// TIA Portal project "Canarias Skills" (V17)
// Prueba de periferia descentralizada ET 200SP

(* hardware
DEVICE "S7-1200 station_1"  S7-1200 Station
   slot 0: "Rack_0"  S7-1200 Rack  Rack  V1.0
   slot 1: "PLC"  CPU 1215C AC/DC/Rly  6ES7 215-1BG40-0XB0  V4.5
DEVICE "GSD device_1"  GSD.Device.PN
   slot 0: "Rack"  Rack  V1.0
   slot 0: "MASTER IO-Link"  AL1100  AL1100
      slot 0: "AL1100"  AL1100
      slot 1: "X1"  X1
         slot 1: "Port 1"  Port 1
         slot 2: "Port 2"  Port 2
      slot 1: "4 Ports_1"  4 Ports  AL1100
         slot 0: "IO-Link Master"  IO-Link Master
   slot 1: "Encoder"  IO-Link In  2 Byte + PQI
   slot 2: "PE"  Digital Input + PQI
   slot 3: "Capacitivo"  Digital Input + PQI
   slot 4: "Disabled_1"  Disabled
DEVICE "SINAMICS G_1"  Sinamics.Device
   slot 0: "	_0"  Rail  SinamicsG120SVecto
   slot 0: "DRIVE_cinta"  G120 CU250S-2 PN Vector  6SL3246-0BA22-1FA0  4.6
      slot 1: "PROFINET interface"  MDD-SinamicsG120-P
   slot 3: "PM240-2 IP20"  PM240-2 IP20  6SL3210-1PB13-8ULx  -
DEVICE "ET 200SP station_1"  ET 200SP-Station
   slot 0: "Rack_0"  Rack  6ES5 710-8MAx1
   slot 0: "IO device_1"  IM 155-6 PN HF  6ES7 155-6AU00-0CN0  V3.1
   slot 1: "DI 8x24VDC HF_1"  DI 8x24VDC HF  6ES7 131-6BF00-0CA0  V1.2
      slot 1: "DI 8x24VDC HF_1"  DI 8x24VDC HF
   slot 2: "DQ 8x24VDC/0.5A HF_1"  DQ 8x24VDC/0.5A HF  6ES7 132-6BF00-0CA0  V1.2
      slot 1: "DQ 8x24VDC/0.5A HF_1"  DQ 8x24VDC/0.5A HF
   slot 3: "Server module_1"  Server module  6ES7 193-6PA00-0AA0  V1.1
      slot 1: "Server module_1"  Server module
   slot 127: "BA 2xRJ45"  BA 2xRJ45  6ES7 193-6AR00-0AA0  V0.0
      slot 1: "Port_1"  X1 P1 R  6ES7 193-6AR00-0AA0  V0.0
      slot 2: "Port_2"  X1 P2 R  6ES7 193-6AR00-0AA0  V0.0
DEVICE "HMI"  KTP700 Basic PN
   slot 0: "HMI"  KTP700 Basic PN  6AV2 123-2GB03-0AX0  17.0.0.0
   slot 1: "HMI_RT_1"  KTP700 Basic PN  6AV2 123-2GB03-0AX0  17.0.0.0
   slot 5: "HMI.IE_CP_1"  PROFINET Interface  17.0.0.0
      slot 1: "PROFINET Interface_1"  PROFINET Interface
         slot 1: "Port_1"  Port
*)

// ===== PLC "PLC"  CPU 1215C AC/DC/Rly =====

VAR_GLOBAL   // PLC tag table "Default tag table"
   "System_Byte" AT %MB1 : Byte;
   "FirstScan" AT %M1.0 : Bool;
   "DiagStatusUpdate" AT %M1.1 : Bool;
   "AlwaysTRUE" AT %M1.2 : Bool;
   "AlwaysFALSE" AT %M1.3 : Bool;
   "Clock_Byte" AT %MB0 : Byte;
   "Clock_10Hz" AT %M0.0 : Bool;
   "Clock_5Hz" AT %M0.1 : Bool;
   "Clock_2.5Hz" AT %M0.2 : Bool;
   "Clock_2Hz" AT %M0.3 : Bool;
   "Clock_1.25Hz" AT %M0.4 : Bool;
   "Clock_1Hz" AT %M0.5 : Bool;
   "Clock_0.625Hz" AT %M0.6 : Bool;
   "Clock_0.5Hz" AT %M0.7 : Bool;
   "Tag_1" AT %Q256.7 : Bool;
   "Tag_2" AT %Q257.7 : Bool;
   "Tag_3" AT %I0.0 : Bool;
   "Tag_4" AT %Q0.0 : Bool;
   "Tag_5" AT %M100.0 : Bool;
END_VAR

VAR_GLOBAL   // PLC tag table "Tag table_1"
   "Encoder" AT %IW68 : Word;
   "Envase" AT %I2.0 : Bool;
   "Llenador_retroceder" AT %Q2.0 : Bool;
   "Llenador_avanzar" AT %Q2.2 : Bool;
   "Cargar_tapa_retroceder" AT %Q2.4 : Bool;
   "Cargar_tapa_avanzar" AT %Q2.6 : Bool;
   "Taponador_retroceder" AT %Q2.1 : Bool;
   "Taponador_avanzar" AT %Q2.5 : Bool;
   "Cargar_tapa_atras" AT %I3.0 : Bool;
   "Cargar_tapa_adelante" AT %I3.1 : Bool;
   "Taponador_atras" AT %I3.2 : Bool;
   "Taponador_adelante" AT %I3.3 : Bool;
   "Mando_driver_cinta" AT %QW256 : Word;
   "Consigna_driver_cinta" AT %QW258 : Word;
   "Estado_driver_cinta" AT %IW256 : Word;
   "Velocidad_cinta" AT %IW258 : Word;
   "R_distancia" AT %M210.0 : Bool;   // Borrar el contador de distancia de la cinta
   "PV_distancia" AT %MW212 : Word;   // Distancia que debe avanzar la cinta
   "Pulso_encoder" AT %I69.0 : Bool;   // Los pulsos del encoder marcan el avance de la cinta
   "PE" AT %I4.1 : Bool;   // Paro de energencia NC
   "CV_distancia" AT %MW214 : Word;   // Distancia que ha recorrido la cinta
   "Q_distancia" AT %M210.1 : Bool;   // Indica que la cinta recorrió la distancia programada
   "Alarmas" AT %MW100 : Word;   // Bits de alarma del HMI
   "ACK_alarmas" AT %MW102 : Word;   // Bits de reconocimiento de alarmas
END_VAR

DATA_BLOCK "Modbus Connect"   // DB1
{ S7_Optimized_Access := 'FALSE' }
VERSION : 0.1
   VAR
      Arduino_1 : Struct
         Configuration : TCON_IP_v4;
         Status : Word;
      END_STRUCT;
   END_VAR
BEGIN
   Arduino_1.Configuration.InterfaceId := 64;
   Arduino_1.Configuration.ID := 16#1;
   Arduino_1.Configuration.ActiveEstablished := TRUE;
   Arduino_1.Configuration.RemoteAddress.ADDR[4] := 200;
   Arduino_1.Configuration.RemoteAddress.ADDR[3] := 0;
   Arduino_1.Configuration.RemoteAddress.ADDR[2] := 168;
   Arduino_1.Configuration.RemoteAddress.ADDR[1] := 192;
   Arduino_1.Configuration.RemotePort := 502;
   Arduino_1.Configuration.LocalPort := 0;
END_DATA_BLOCK

DATA_BLOCK "Modbus Buffer"   // DB3
{ S7_Optimized_Access := 'FALSE' }
VERSION : 0.1
   VAR
      Datos : Array[0..100] of Word;
   END_VAR
BEGIN
END_DATA_BLOCK

DATA_BLOCK "Modo_automatico_DB"   // DB4
{ S7_Optimized_Access := 'TRUE' }
VERSION : 0.1
// stored: InstanceOfName Modo_automatico
"Modo_automatico"
BEGIN
END_DATA_BLOCK

DATA_BLOCK "Datos_maquina"   // DB5
{ S7_Optimized_Access := 'TRUE' }
VERSION : 0.1
   VAR RETAIN
      pp_mm : Int := 2;   // Pulsos de encoder por cada milímetro de avance de cinta
      Desviador_bloquear : Word := 0;   // Posición del desviador para bloquear pieza
      Desviador_rechazar : Word := 37;   // Posición del desviador para rechazar pieza
      Desviador_aceptar : Word := 82;   // Posición del desviador para aceptar pieza
      Distancia_inspeccion : Word := 50;   // Distancia en mm hasta el inspector
      Distancia_desviador : Word := 100;   // Distancia en mm hasta el desviador
      Distancia_llenadora : Word := 200;   // Distancia en mm hasta la llenadora
      Distancia_taponadora : Word := 300;   // Distancia en mm hasta la taponadora
      Distancia_salida : Word := 400;   // Distancia en mm hasta la salida de la cinta
      Cinta_en_espera : Word := 16#047E;   // Driver cinta listo y en espera
      Cinta_en_marcha : Word := 16#0C7F;   // Driver cinta en avance
      Consigna_cinta : Int := 8000;   // Consigna de velocidad de la cinta
      Freno_en_cinta : Word := 16#043F;   // Activar freno con rampa driver cinta
      Freno_en_cinta_rapido : Word := 16#043D;   // Activar freno rápìdo driver cinta
      Total_envasados : Word;   // Catidad de envases producidos
      Total_rechazados : Word;   // Cantidad de envases rechazados
   END_VAR
   VAR
      HMI_llenador_retroceder : Bool;   // Lo que sigue son maniobras en modo manual desde el HMI
      HMI_llenador_avanzar : Bool;
      HMI_cargar_tapa_retroceder : Bool;
      HMI_cargar_tapa_avanzar : Bool;
      HMI_taponar_retroceder : Bool;
      HMI_taponar_avanzar : Bool;
      HMI_desviador_bloquear : Bool;
      HMI_desviador_rechazar : Bool;
      HMI_desviador_aceptar : Bool;
      HMI_driver_listo : Bool;
      HMI_driver_acusar_fallo : Bool;   // Manobras en modo manual de la cinta
      HMI_driver_detener_rampa : Bool;
      HMI_driver_detener_freno : Bool;
      HMI_driver_marcha : Bool;
      HMI_marcha : Bool;   // Marcha desde el HMI
      HMI_paro : Bool;   // Paro desde el HMI
      HMI_reset : Bool;   // Reset desde el HMI
   END_VAR
   VAR RETAIN
      HMI_manual_automatico : Bool;   // Modo de operación desde el HMI
      Estado : Struct
         Esperando_marcha : Bool;
         En_marcha : Bool;
         En_paro : Bool;
         En_PE : Bool;
         Esperando_reset : Bool;
      END_STRUCT;
   END_VAR
   VAR
      Inspector : Struct
         Enviar : Bool;
         Recibir : Bool;
         Recibido_ok : Bool;
         Recibido_error : Bool;
      END_STRUCT;
   END_VAR
BEGIN
END_DATA_BLOCK

DATA_BLOCK "Paro_emergencia_DB"   // DB10
{ S7_Optimized_Access := 'TRUE' }
VERSION : 0.1
// stored: InstanceOfName Paro_emergencia
"Paro_emergencia"
BEGIN
END_DATA_BLOCK

DATA_BLOCK "Raspberry PI Buffer"   // DB13
{ S7_Optimized_Access := 'FALSE' }
VERSION : 0.1
   VAR
      Data_send : Array[0..100] of Char;
      Data_rcv : Array[0..29] of Char;
   END_VAR
BEGIN
   Data_send[9] := '"';
   Data_send[8] := 'd';
   Data_send[7] := 'n';
   Data_send[6] := 'a';
   Data_send[5] := 'm';
   Data_send[4] := 'm';
   Data_send[3] := 'o';
   Data_send[2] := 'c';
   Data_send[1] := '"';
   Data_send[0] := '{';
   Data_send[10] := ':';   // {Command=I} para inferir objeto
   Data_send[11] := '"';
   Data_send[12] := 'I';
   Data_send[13] := '"';
   Data_send[14] := '}';
END_DATA_BLOCK

// folder: System blocks/Program resources

DATA_BLOCK "Distancia"   // DB6
{ S7_Optimized_Access := 'TRUE' }
AUTHOR : Simatic
FAMILY : IEC
NAME : CNTR
VERSION : 1.0
// stored: InstanceOfName IEC_COUNTER
"IEC_COUNTER"
BEGIN
END_DATA_BLOCK

DATA_BLOCK "IEC_Timer_0_DB"   // DB7
{ S7_Optimized_Access := 'TRUE' }
AUTHOR : Simatic
FAMILY : IEC
NAME : IEC_TMR
VERSION : 1.0
// stored: InstanceOfName IEC_TIMER
"IEC_TIMER"
BEGIN
END_DATA_BLOCK

DATA_BLOCK "IEC_Timer_0_DB_1"   // DB8
{ S7_Optimized_Access := 'TRUE' }
AUTHOR : Simatic
FAMILY : IEC
NAME : IEC_TMR
VERSION : 1.0
// stored: InstanceOfName IEC_TIMER
"IEC_TIMER"
BEGIN
END_DATA_BLOCK

DATA_BLOCK "IEC_Timer_0_DB_2"   // DB9
{ S7_Optimized_Access := 'TRUE' }
AUTHOR : Simatic
FAMILY : IEC
NAME : IEC_TMR
VERSION : 1.0
// stored: InstanceOfName IEC_TIMER
"IEC_TIMER"
BEGIN
END_DATA_BLOCK

DATA_BLOCK "IEC_Timer_0_DB_3"   // DB11
{ S7_Optimized_Access := 'TRUE' }
AUTHOR : Simatic
FAMILY : IEC
NAME : IEC_TMR
VERSION : 1.0
// stored: InstanceOfName IEC_TIMER
"IEC_TIMER"
BEGIN
END_DATA_BLOCK

DATA_BLOCK "PLC_Receive_DB"   // DB15
{ S7_Optimized_Access := 'TRUE' }
AUTHOR : SIMATIC
FAMILY : MC7Plus
NAME : TC_IP_v4
VERSION : 1.0
// stored: InstanceOfName TCON_IP_v4
"TCON_IP_v4"
BEGIN
   ID := 3;
   InterfaceId := 64;
   LocalPort := 2000;
   RemotePort := 2000;
   ActiveEstablished := true;
   RemoteAddress.ADDR[1] := 192;
   RemoteAddress.ADDR[2] := 168;
   RemoteAddress.ADDR[4] := 241;
END_DATA_BLOCK

DATA_BLOCK "IEC_Timer_0_DB_4"   // DB16
{ S7_Optimized_Access := 'TRUE' }
AUTHOR : Simatic
FAMILY : IEC
NAME : IEC_TMR
VERSION : 1.0
// stored: InstanceOfName IEC_TIMER
"IEC_TIMER"
BEGIN
END_DATA_BLOCK

DATA_BLOCK "IEC_Timer_0_DB_5"   // DB17
{ S7_Optimized_Access := 'TRUE' }
AUTHOR : Simatic
FAMILY : IEC
NAME : IEC_TMR
VERSION : 1.0
// stored: InstanceOfName IEC_TIMER
"IEC_TIMER"
BEGIN
END_DATA_BLOCK

DATA_BLOCK "IEC_Timer_0_DB_6"   // DB18
{ S7_Optimized_Access := 'TRUE' }
AUTHOR : Simatic
FAMILY : IEC
NAME : IEC_TMR
VERSION : 1.0
// stored: InstanceOfName IEC_TIMER
"IEC_TIMER"
BEGIN
END_DATA_BLOCK

DATA_BLOCK "IEC_Timer_0_DB_7"   // DB19
{ S7_Optimized_Access := 'TRUE' }
AUTHOR : Simatic
FAMILY : IEC
NAME : IEC_TMR
VERSION : 1.0
// stored: InstanceOfName IEC_TIMER
"IEC_TIMER"
BEGIN
END_DATA_BLOCK

// folder: (top level)

FUNCTION_BLOCK "Paro_emergencia"   // FB1, LAD
{ S7_Optimized_Access := 'TRUE' }
VERSION : 0.1
   VAR
      Etapa_0 : Bool := true;
      Etapa_1 : Bool;
      Etapa_2 : Bool;
   END_VAR
   VAR_TEMP   // added for the SCL form of the ladder/FBD networks
      _w1 : Bool;
   END_VAR
BEGIN

REGION Network 1: Emergencia Etapa 0
   // - Activar marca de situación de Paro de Emergencia
   // - Desactivar todos los distribuidores neumáticos
   // - Detener cinta con freno
   // - Desviador a posición de aceptar envase
   // - Reset contador de distancia de cinta
   // 
   // Esperar la desactivación del Paro de Emergencia (PE) y la pulsación de Reset en el HMI
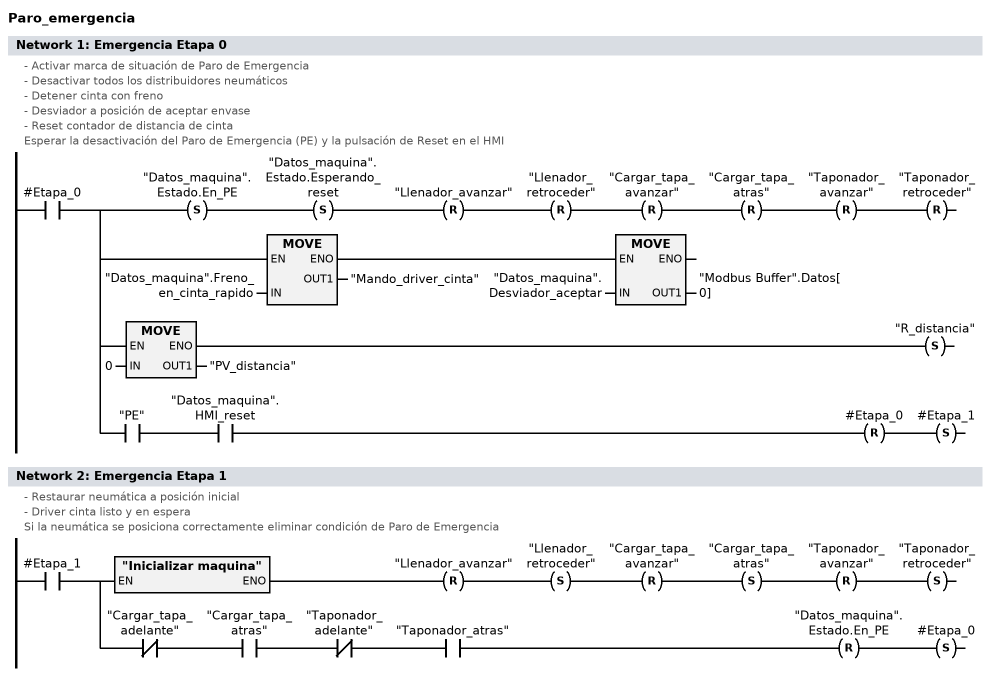
   RUNG wire#powerrail
      Contact( #Etapa_0 )
      wire#w1
      S_Coil( "Datos_maquina".Estado.En_PE )
      S_Coil( "Datos_maquina".Estado.Esperando_reset )
      R_Coil( "Llenador_avanzar" )
      R_Coil( "Llenador_retroceder" )
      R_Coil( "Cargar_tapa_avanzar" )
      R_Coil( "Cargar_tapa_atras" )
      R_Coil( "Taponador_avanzar" )
      R_Coil( "Taponador_retroceder" )
   END_RUNG
   RUNG wire#w1
      Move(in := "Datos_maquina".Freno_en_cinta_rapido, out1 => "Mando_driver_cinta")
      Move(in := "Datos_maquina".Desviador_aceptar, out1 => "Modbus Buffer".Datos[0])
   END_RUNG
   RUNG wire#w1
      Move(in := 0, out1 => "PV_distancia")
      S_Coil( "R_distancia" )
   END_RUNG
   RUNG wire#w1
      Contact( "PE" )
      Contact( "Datos_maquina".HMI_reset )
      R_Coil( #Etapa_0 )
      S_Coil( #Etapa_1 )
   END_RUNG
   // the same network as SCL:
   IF #Etapa_0 THEN
       "Datos_maquina".Estado.En_PE := TRUE;
       "Datos_maquina".Estado.Esperando_reset := TRUE;
       "Llenador_avanzar" := FALSE;
       "Llenador_retroceder" := FALSE;
       "Cargar_tapa_avanzar" := FALSE;
       "Cargar_tapa_atras" := FALSE;
       "Taponador_avanzar" := FALSE;
       "Taponador_retroceder" := FALSE;
       "Mando_driver_cinta" := "Datos_maquina".Freno_en_cinta_rapido;
       "Modbus Buffer".Datos[0] := "Datos_maquina".Desviador_aceptar;
       "PV_distancia" := 0;
       "R_distancia" := TRUE;
   END_IF;
   #_w1 := #Etapa_0 AND "PE" AND "Datos_maquina".HMI_reset;
   IF #_w1 THEN
       #Etapa_0 := FALSE;
       #Etapa_1 := TRUE;
   END_IF;
END_REGION

REGION Network 2: Emergencia Etapa 1
   // - Restaurar neumática a posición inicial
   // - Driver cinta listo y en espera
   // 
   // Si la neumática se posiciona correctamente eliminar condición de Paro de Emergencia
   RUNG wire#powerrail
      Contact( #Etapa_1 )
      wire#w1
      "Inicializar maquina"()
      R_Coil( "Llenador_avanzar" )
      S_Coil( "Llenador_retroceder" )
      R_Coil( "Cargar_tapa_avanzar" )
      S_Coil( "Cargar_tapa_atras" )
      R_Coil( "Taponador_avanzar" )
      S_Coil( "Taponador_retroceder" )
   END_RUNG
   RUNG wire#w1
      I_Contact( "Cargar_tapa_adelante" )
      Contact( "Cargar_tapa_atras" )
      I_Contact( "Taponador_adelante" )
      Contact( "Taponador_atras" )
      R_Coil( "Datos_maquina".Estado.En_PE )
      S_Coil( #Etapa_0 )
   END_RUNG
   // the same network as SCL:
   "Inicializar maquina"(EN := #Etapa_1, ENO => #_w1);
   IF #_w1 THEN
       "Llenador_avanzar" := FALSE;
       "Llenador_retroceder" := TRUE;
       "Cargar_tapa_avanzar" := FALSE;
       "Cargar_tapa_atras" := TRUE;
       "Taponador_avanzar" := FALSE;
       "Taponador_retroceder" := TRUE;
   END_IF;
   IF #Etapa_1 AND NOT "Cargar_tapa_adelante" AND "Cargar_tapa_atras" AND NOT "Taponador_adelante" AND "Taponador_atras" THEN
       "Datos_maquina".Estado.En_PE := FALSE;
       #Etapa_0 := TRUE;
   END_IF;
END_REGION
END_FUNCTION_BLOCK

FUNCTION_BLOCK "Modo_automatico"   // FB2, LAD
{ S7_Optimized_Access := 'TRUE' }
VERSION : 0.1
   VAR
      Etapa_0 : Bool := true;
      Etapa_1 : Bool;
      Etapa_2 : Bool;
      Etapa_3 : Bool;
      Etapa_4 : Bool;
      Etapa_5 : Bool;
      Etapa_6 : Bool;
      Etapa_7 : Bool;
      Etapa_8 : Bool;
      Etapa_9 : Bool;
      Etapa_10 : Bool;
      Etapa_11 : Bool;
      Etapa_12 : Bool;
      Etapa_13 : Bool;
      Aux1 : Bool;   // Para detectar flanco postivo del HMI_paro
   END_VAR
   VAR_TEMP
      Resultado : String;
   END_VAR
   VAR_TEMP   // added for the SCL form of the ladder/FBD networks
      _w1 : Bool;
      _w2 : Bool;
   END_VAR
BEGIN

REGION Network 1: Maniobra de Paro
   // - Detiene la cinta
   // - Deesactiva todas las etapas del GRAFCET
   // - Espera un rearme desde HMI para situarse en la etapa 0 del GRAFCET
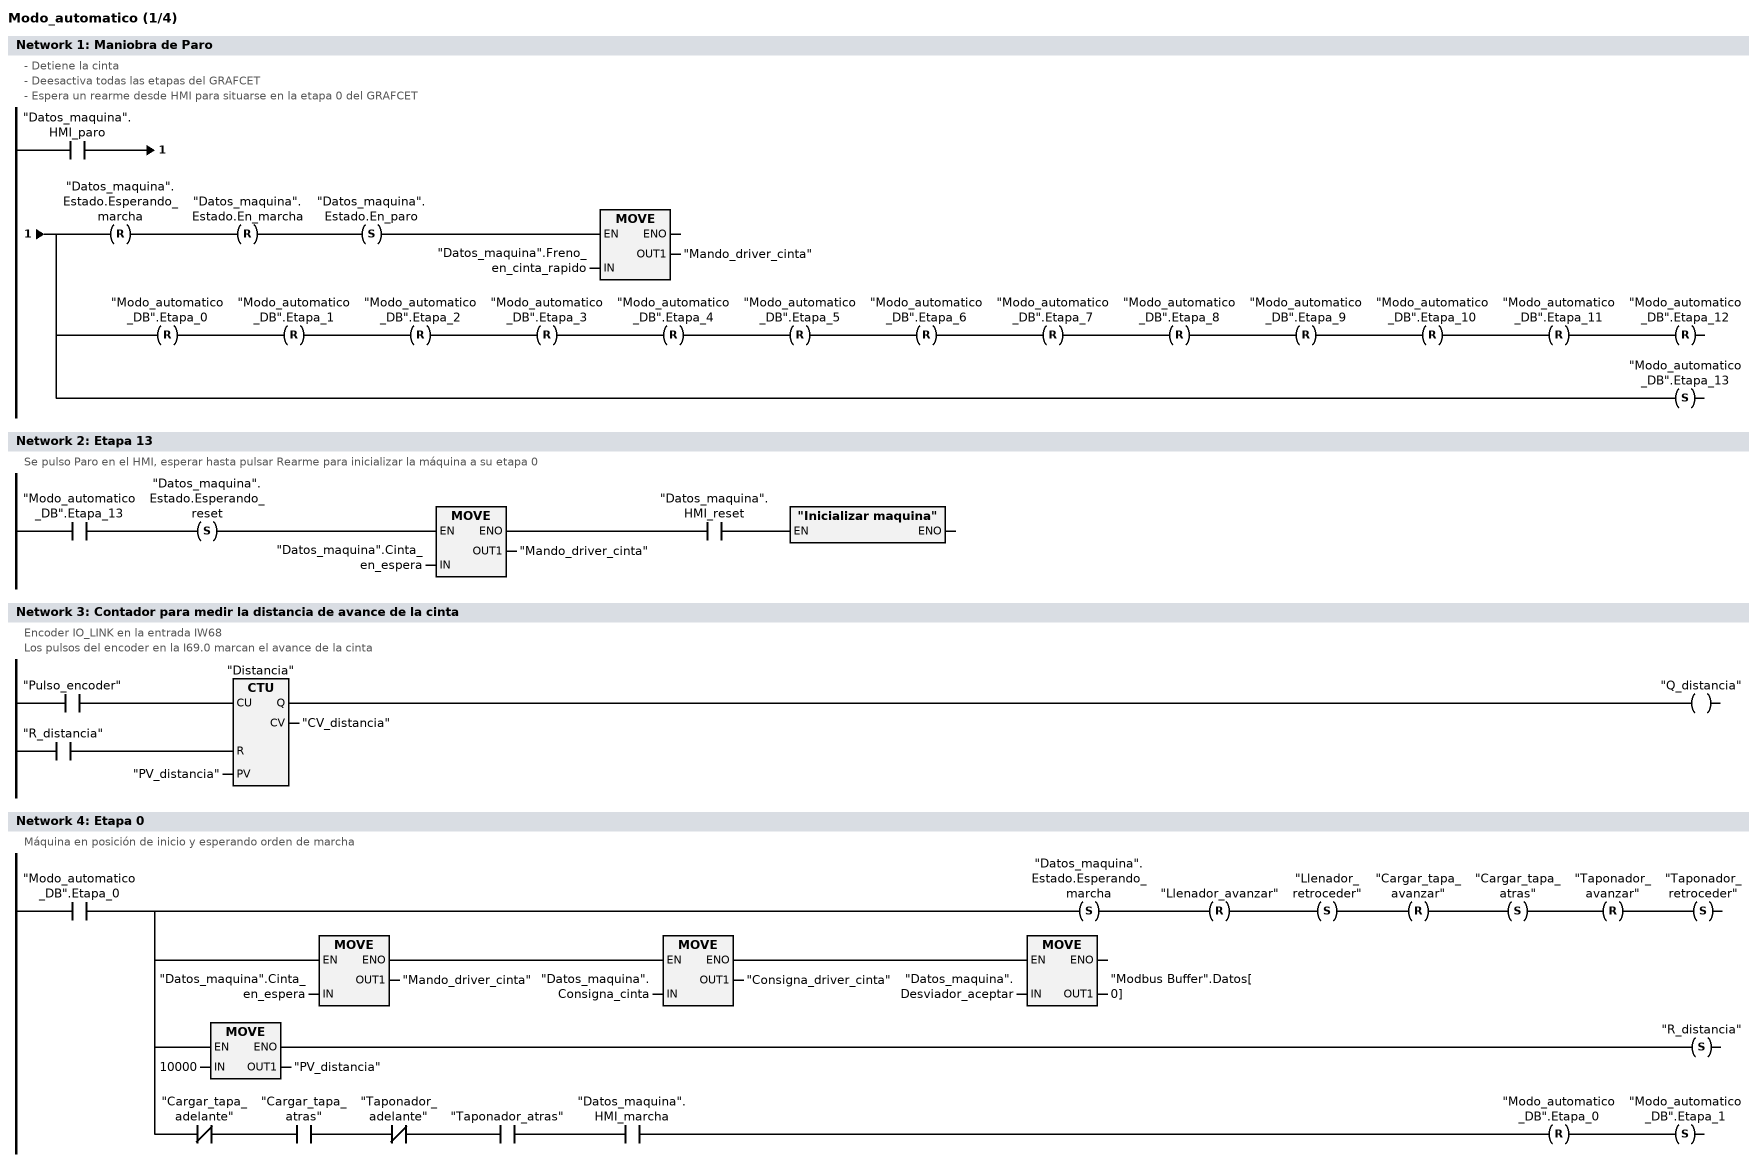
   RUNG wire#powerrail
      Contact( "Datos_maquina".HMI_paro )
      wire#w1
      R_Coil( "Datos_maquina".Estado.Esperando_marcha )
      R_Coil( "Datos_maquina".Estado.En_marcha )
      S_Coil( "Datos_maquina".Estado.En_paro )
      Move(in := "Datos_maquina".Freno_en_cinta_rapido, out1 => "Mando_driver_cinta")
   END_RUNG
   RUNG wire#w1
      R_Coil( "Modo_automatico_DB".Etapa_0 )
      R_Coil( "Modo_automatico_DB".Etapa_1 )
      R_Coil( "Modo_automatico_DB".Etapa_2 )
      R_Coil( "Modo_automatico_DB".Etapa_3 )
      R_Coil( "Modo_automatico_DB".Etapa_4 )
      R_Coil( "Modo_automatico_DB".Etapa_5 )
      R_Coil( "Modo_automatico_DB".Etapa_6 )
      R_Coil( "Modo_automatico_DB".Etapa_7 )
      R_Coil( "Modo_automatico_DB".Etapa_8 )
      R_Coil( "Modo_automatico_DB".Etapa_9 )
      R_Coil( "Modo_automatico_DB".Etapa_10 )
      R_Coil( "Modo_automatico_DB".Etapa_11 )
      R_Coil( "Modo_automatico_DB".Etapa_12 )
   END_RUNG
   RUNG wire#w1
      S_Coil( "Modo_automatico_DB".Etapa_13 )
   END_RUNG
   // the same network as SCL:
   IF "Datos_maquina".HMI_paro THEN
       "Datos_maquina".Estado.Esperando_marcha := FALSE;
       "Datos_maquina".Estado.En_marcha := FALSE;
       "Datos_maquina".Estado.En_paro := TRUE;
       "Mando_driver_cinta" := "Datos_maquina".Freno_en_cinta_rapido;
       "Modo_automatico_DB".Etapa_0 := FALSE;
       "Modo_automatico_DB".Etapa_1 := FALSE;
       "Modo_automatico_DB".Etapa_2 := FALSE;
       "Modo_automatico_DB".Etapa_3 := FALSE;
       "Modo_automatico_DB".Etapa_4 := FALSE;
       "Modo_automatico_DB".Etapa_5 := FALSE;
       "Modo_automatico_DB".Etapa_6 := FALSE;
       "Modo_automatico_DB".Etapa_7 := FALSE;
       "Modo_automatico_DB".Etapa_8 := FALSE;
       "Modo_automatico_DB".Etapa_9 := FALSE;
       "Modo_automatico_DB".Etapa_10 := FALSE;
       "Modo_automatico_DB".Etapa_11 := FALSE;
       "Modo_automatico_DB".Etapa_12 := FALSE;
       "Modo_automatico_DB".Etapa_13 := TRUE;
   END_IF;
END_REGION

REGION Network 2: Etapa 13
   // Se pulso Paro en el HMI, esperar hasta pulsar Rearme para inicializar la máquina a su etapa 0
   RUNG wire#powerrail
      Contact( "Modo_automatico_DB".Etapa_13 )
      S_Coil( "Datos_maquina".Estado.Esperando_reset )
      Move(in := "Datos_maquina".Cinta_en_espera, out1 => "Mando_driver_cinta")
      Contact( "Datos_maquina".HMI_reset )
      "Inicializar maquina"()
   END_RUNG
   // the same network as SCL:
   IF "Modo_automatico_DB".Etapa_13 THEN
       "Datos_maquina".Estado.Esperando_reset := TRUE;
       "Mando_driver_cinta" := "Datos_maquina".Cinta_en_espera;
   END_IF;
   IF "Modo_automatico_DB".Etapa_13 AND "Datos_maquina".HMI_reset THEN "Inicializar maquina"(); END_IF;
END_REGION

REGION Network 3: Contador para medir la distancia de avance de la cinta
   // Encoder IO_LINK en la entrada IW68
   // Los pulsos del encoder en la I69.0 marcan el avance de la cinta
   "Distancia".CTU(CU := "Pulso_encoder", R := "R_distancia", PV := "PV_distancia", CV => "CV_distancia");
   "Q_distancia" := "Distancia".Q;
END_REGION

REGION Network 4: Etapa 0
   // Máquina en posición de inicio y esperando orden de marcha
   RUNG wire#powerrail
      Contact( "Modo_automatico_DB".Etapa_0 )
      wire#w1
      S_Coil( "Datos_maquina".Estado.Esperando_marcha )
      R_Coil( "Llenador_avanzar" )
      S_Coil( "Llenador_retroceder" )
      R_Coil( "Cargar_tapa_avanzar" )
      S_Coil( "Cargar_tapa_atras" )
      R_Coil( "Taponador_avanzar" )
      S_Coil( "Taponador_retroceder" )
   END_RUNG
   RUNG wire#w1
      Move(in := "Datos_maquina".Cinta_en_espera, out1 => "Mando_driver_cinta")
      Move(in := "Datos_maquina".Consigna_cinta, out1 => "Consigna_driver_cinta")
      Move(in := "Datos_maquina".Desviador_aceptar, out1 => "Modbus Buffer".Datos[0])
   END_RUNG
   RUNG wire#w1
      Move(in := 10000, out1 => "PV_distancia")
      S_Coil( "R_distancia" )
   END_RUNG
   RUNG wire#w1
      I_Contact( "Cargar_tapa_adelante" )
      Contact( "Cargar_tapa_atras" )
      I_Contact( "Taponador_adelante" )
      Contact( "Taponador_atras" )
      Contact( "Datos_maquina".HMI_marcha )
      R_Coil( "Modo_automatico_DB".Etapa_0 )
      S_Coil( "Modo_automatico_DB".Etapa_1 )
   END_RUNG
   // the same network as SCL:
   IF "Modo_automatico_DB".Etapa_0 THEN
       "Datos_maquina".Estado.Esperando_marcha := TRUE;
       "Llenador_avanzar" := FALSE;
       "Llenador_retroceder" := TRUE;
       "Cargar_tapa_avanzar" := FALSE;
       "Cargar_tapa_atras" := TRUE;
       "Taponador_avanzar" := FALSE;
       "Taponador_retroceder" := TRUE;
       "Mando_driver_cinta" := "Datos_maquina".Cinta_en_espera;
       "Consigna_driver_cinta" := "Datos_maquina".Consigna_cinta;
       "Modbus Buffer".Datos[0] := "Datos_maquina".Desviador_aceptar;
       "PV_distancia" := 10000;
       "R_distancia" := TRUE;
   END_IF;
   #_w1 := "Modo_automatico_DB".Etapa_0 AND NOT "Cargar_tapa_adelante" AND "Cargar_tapa_atras" AND NOT "Taponador_adelante" AND "Taponador_atras" AND "Datos_maquina".HMI_marcha;
   IF #_w1 THEN
       "Modo_automatico_DB".Etapa_0 := FALSE;
       "Modo_automatico_DB".Etapa_1 := TRUE;
   END_IF;
END_REGION

REGION Network 5: Etapa 1
   // Probar desviador a bloquear pieza
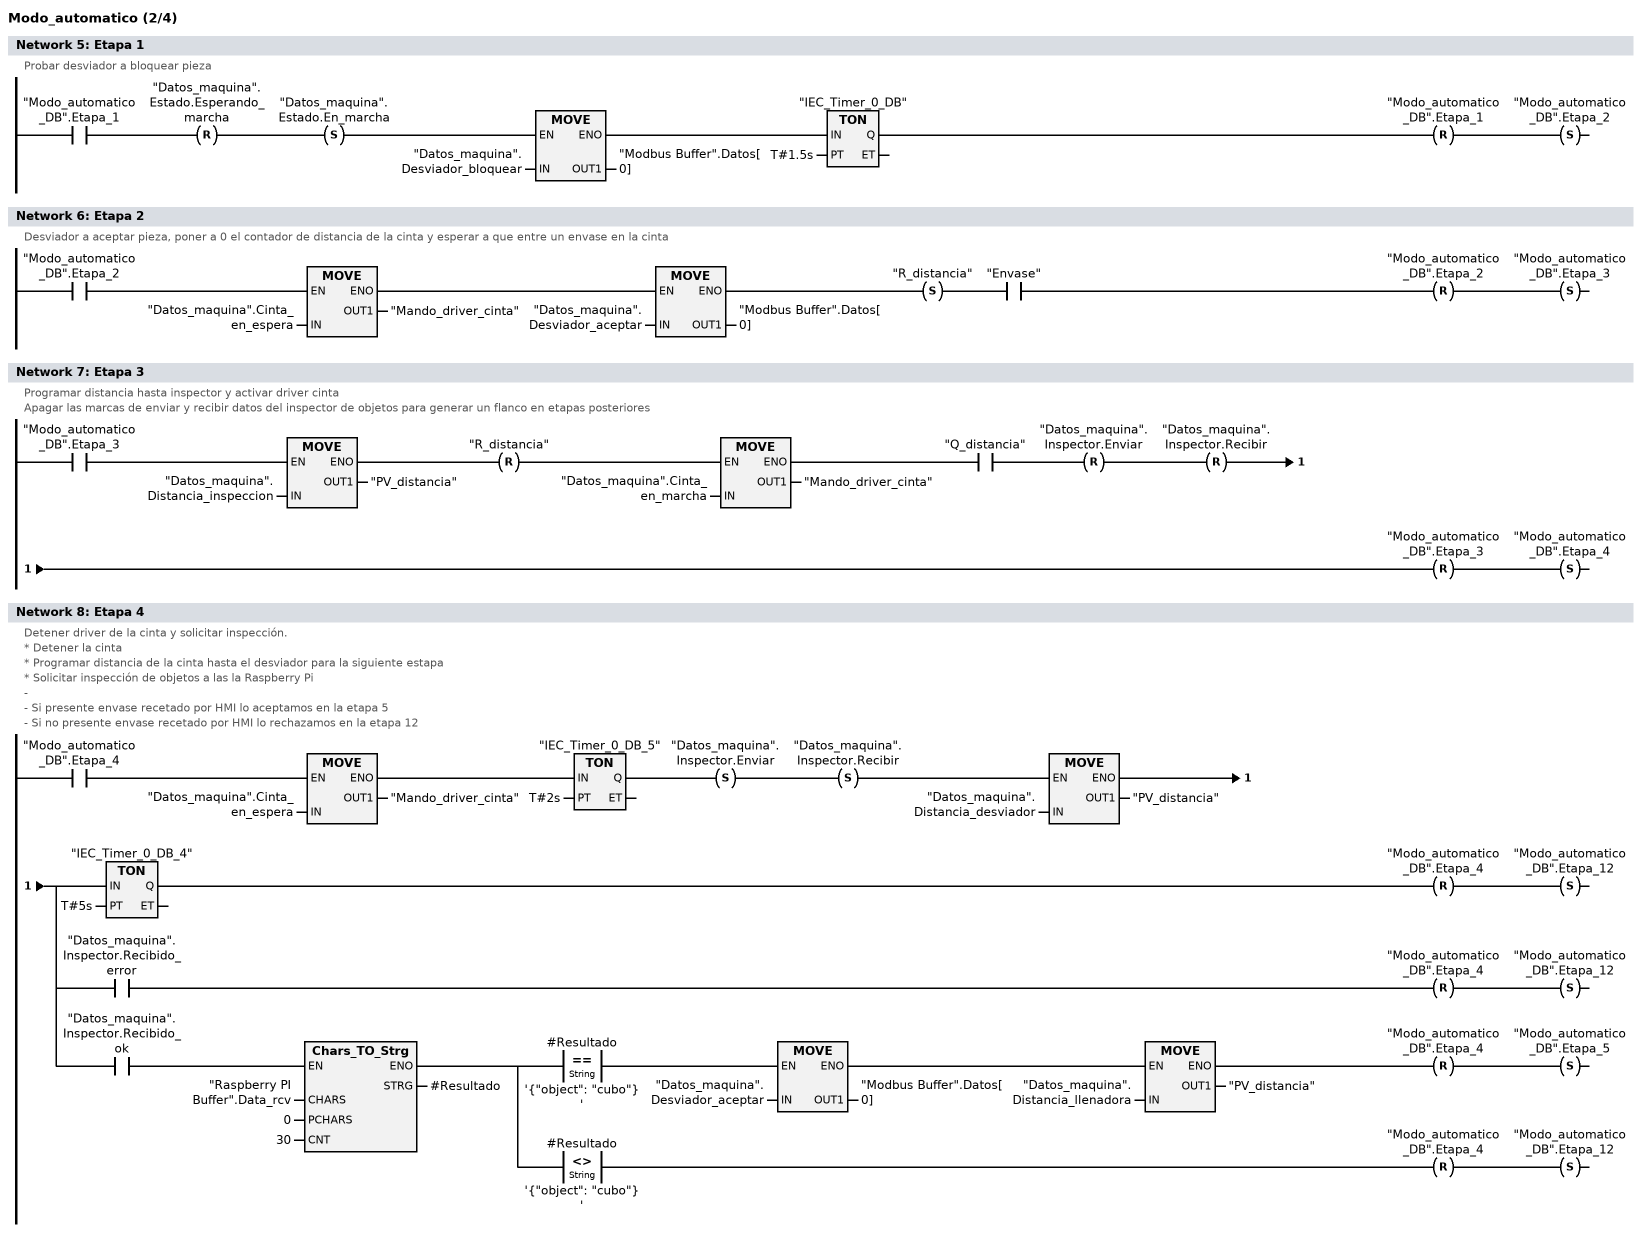
   IF "Modo_automatico_DB".Etapa_1 THEN
       "Datos_maquina".Estado.Esperando_marcha := FALSE;
       "Datos_maquina".Estado.En_marcha := TRUE;
       "Modbus Buffer".Datos[0] := "Datos_maquina".Desviador_bloquear;
   END_IF;
   "IEC_Timer_0_DB".TON(IN := "Modo_automatico_DB".Etapa_1, PT := T#1.5s);
   IF "IEC_Timer_0_DB".Q THEN
       "Modo_automatico_DB".Etapa_1 := FALSE;
       "Modo_automatico_DB".Etapa_2 := TRUE;
   END_IF;
END_REGION

REGION Network 6: Etapa 2
   // Desviador a aceptar pieza, poner a 0 el contador de distancia de la cinta y esperar a que entre un envase en la cinta
   RUNG wire#powerrail
      Contact( "Modo_automatico_DB".Etapa_2 )
      Move(in := "Datos_maquina".Cinta_en_espera, out1 => "Mando_driver_cinta")
      Move(in := "Datos_maquina".Desviador_aceptar, out1 => "Modbus Buffer".Datos[0])
      S_Coil( "R_distancia" )
      Contact( "Envase" )
      R_Coil( "Modo_automatico_DB".Etapa_2 )
      S_Coil( "Modo_automatico_DB".Etapa_3 )
   END_RUNG
   // the same network as SCL:
   IF "Modo_automatico_DB".Etapa_2 THEN
       "Mando_driver_cinta" := "Datos_maquina".Cinta_en_espera;
       "Modbus Buffer".Datos[0] := "Datos_maquina".Desviador_aceptar;
       "R_distancia" := TRUE;
   END_IF;
   #_w1 := "Modo_automatico_DB".Etapa_2 AND "Envase";
   IF #_w1 THEN
       "Modo_automatico_DB".Etapa_2 := FALSE;
       "Modo_automatico_DB".Etapa_3 := TRUE;
   END_IF;
END_REGION

REGION Network 7: Etapa 3
   // Programar distancia hasta inspector y activar driver cinta 
   // Apagar las marcas de enviar y recibir datos del inspector de objetos para generar un flanco en etapas posteriores
   RUNG wire#powerrail
      Contact( "Modo_automatico_DB".Etapa_3 )
      Move(in := "Datos_maquina".Distancia_inspeccion, out1 => "PV_distancia")
      R_Coil( "R_distancia" )
      Move(in := "Datos_maquina".Cinta_en_marcha, out1 => "Mando_driver_cinta")
      Contact( "Q_distancia" )
      R_Coil( "Datos_maquina".Inspector.Enviar )
      R_Coil( "Datos_maquina".Inspector.Recibir )
      R_Coil( "Modo_automatico_DB".Etapa_3 )
      S_Coil( "Modo_automatico_DB".Etapa_4 )
   END_RUNG
   // the same network as SCL:
   IF "Modo_automatico_DB".Etapa_3 THEN
       "PV_distancia" := "Datos_maquina".Distancia_inspeccion;
       "R_distancia" := FALSE;
       "Mando_driver_cinta" := "Datos_maquina".Cinta_en_marcha;
   END_IF;
   IF "Modo_automatico_DB".Etapa_3 AND "Q_distancia" THEN
       "Datos_maquina".Inspector.Enviar := FALSE;
       "Datos_maquina".Inspector.Recibir := FALSE;
   END_IF;
   #_w1 := "Modo_automatico_DB".Etapa_3 AND "Q_distancia";
   IF #_w1 THEN
       "Modo_automatico_DB".Etapa_3 := FALSE;
       "Modo_automatico_DB".Etapa_4 := TRUE;
   END_IF;
END_REGION

REGION Network 8: Etapa 4
   // Detener driver de la cinta y solicitar inspección.
   // 
   // * Detener la cinta
   // * Programar distancia de la cinta hasta el desviador para la siguiente estapa
   // * Solicitar inspección de objetos a las la Raspberry Pi
   //    - 
   //    - Si presente envase recetado por HMI lo aceptamos en la etapa 5
   //    - Si no presente envase recetado por HMI lo rechazamos en la etapa 12
   // no SCL statement known for Chars_TO_Strg: written as a call
   // ENO of a box is taken as its EN; it also drops when the box reports an error
   IF "Modo_automatico_DB".Etapa_4 THEN "Mando_driver_cinta" := "Datos_maquina".Cinta_en_espera; END_IF;
   "IEC_Timer_0_DB_5".TON(IN := "Modo_automatico_DB".Etapa_4, PT := T#2s);
   IF "IEC_Timer_0_DB_5".Q THEN
       "Datos_maquina".Inspector.Enviar := TRUE;
       "Datos_maquina".Inspector.Recibir := TRUE;
       "PV_distancia" := "Datos_maquina".Distancia_desviador;
   END_IF;
   "IEC_Timer_0_DB_4".TON(IN := "IEC_Timer_0_DB_5".Q, PT := T#5s);
   IF "IEC_Timer_0_DB_4".Q THEN
       "Modo_automatico_DB".Etapa_4 := FALSE;
       "Modo_automatico_DB".Etapa_12 := TRUE;
   END_IF;
   IF "IEC_Timer_0_DB_5".Q AND "Datos_maquina".Inspector.Recibido_error THEN
       "Modo_automatico_DB".Etapa_4 := FALSE;
       "Modo_automatico_DB".Etapa_12 := TRUE;
   END_IF;
   #_w1 := "IEC_Timer_0_DB_5".Q AND "Datos_maquina".Inspector.Recibido_ok;
   IF #_w1 THEN
       Chars_TO_Strg(Chars := "Raspberry PI Buffer".Data_rcv, pChars := 0, Cnt := 30, Strg => #Resultado);
   END_IF;
   IF #_w1 AND (#Resultado = '{"object": "cubo"}            ') THEN
       "Modbus Buffer".Datos[0] := "Datos_maquina".Desviador_aceptar;
       "PV_distancia" := "Datos_maquina".Distancia_llenadora;
       "Modo_automatico_DB".Etapa_4 := FALSE;
       "Modo_automatico_DB".Etapa_5 := TRUE;
   END_IF;
   IF #_w1 AND (#Resultado <> '{"object": "cubo"}            ') THEN
       "Modo_automatico_DB".Etapa_4 := FALSE;
       "Modo_automatico_DB".Etapa_12 := TRUE;
   END_IF;
END_REGION

REGION Network 9: Etapa 5
   // Aceptar envase y moverlo hasta la llenadora
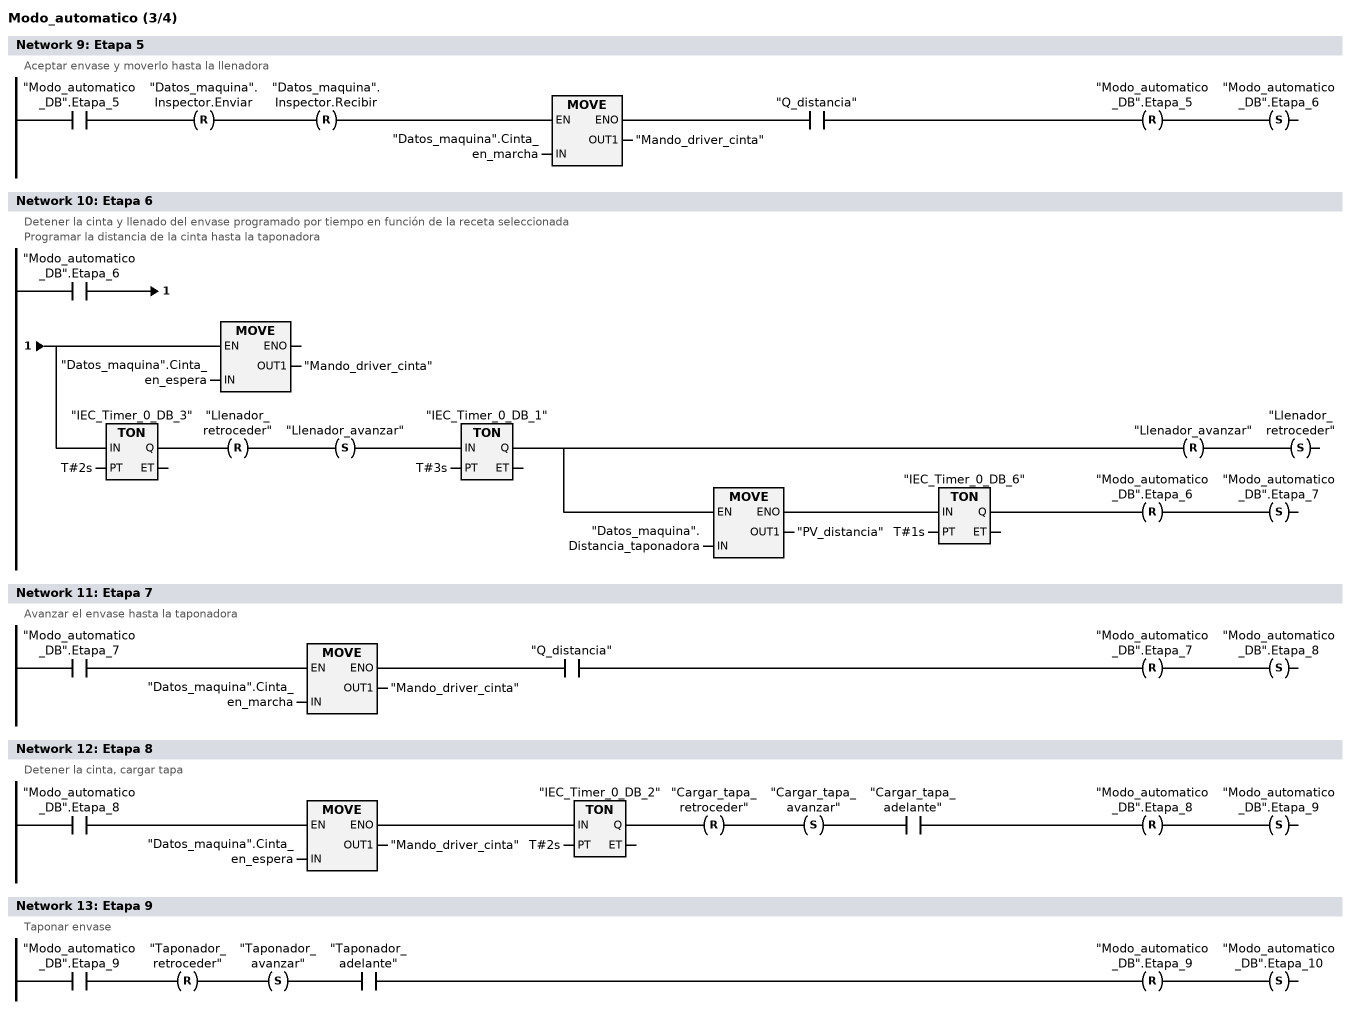
   RUNG wire#powerrail
      Contact( "Modo_automatico_DB".Etapa_5 )
      R_Coil( "Datos_maquina".Inspector.Enviar )
      R_Coil( "Datos_maquina".Inspector.Recibir )
      Move(in := "Datos_maquina".Cinta_en_marcha, out1 => "Mando_driver_cinta")
      Contact( "Q_distancia" )
      R_Coil( "Modo_automatico_DB".Etapa_5 )
      S_Coil( "Modo_automatico_DB".Etapa_6 )
   END_RUNG
   // the same network as SCL:
   IF "Modo_automatico_DB".Etapa_5 THEN
       "Datos_maquina".Inspector.Enviar := FALSE;
       "Datos_maquina".Inspector.Recibir := FALSE;
       "Mando_driver_cinta" := "Datos_maquina".Cinta_en_marcha;
   END_IF;
   #_w1 := "Modo_automatico_DB".Etapa_5 AND "Q_distancia";
   IF #_w1 THEN
       "Modo_automatico_DB".Etapa_5 := FALSE;
       "Modo_automatico_DB".Etapa_6 := TRUE;
   END_IF;
END_REGION

REGION Network 10: Etapa 6
   // Detener la cinta y llenado del envase programado por tiempo en función de la receta seleccionada
   // Programar la distancia de la cinta hasta la taponadora
   IF "Modo_automatico_DB".Etapa_6 THEN "Mando_driver_cinta" := "Datos_maquina".Cinta_en_espera; END_IF;
   "IEC_Timer_0_DB_3".TON(IN := "Modo_automatico_DB".Etapa_6, PT := T#2s);
   IF "IEC_Timer_0_DB_3".Q THEN
       "Llenador_retroceder" := FALSE;
       "Llenador_avanzar" := TRUE;
   END_IF;
   "IEC_Timer_0_DB_1".TON(IN := "IEC_Timer_0_DB_3".Q, PT := T#3s);
   IF "IEC_Timer_0_DB_1".Q THEN
       "Llenador_avanzar" := FALSE;
       "Llenador_retroceder" := TRUE;
       "PV_distancia" := "Datos_maquina".Distancia_taponadora;
   END_IF;
   "IEC_Timer_0_DB_6".TON(IN := "IEC_Timer_0_DB_1".Q, PT := T#1s);
   IF "IEC_Timer_0_DB_6".Q THEN
       "Modo_automatico_DB".Etapa_6 := FALSE;
       "Modo_automatico_DB".Etapa_7 := TRUE;
   END_IF;
END_REGION

REGION Network 11: Etapa 7
   // Avanzar el envase hasta la taponadora
   RUNG wire#powerrail
      Contact( "Modo_automatico_DB".Etapa_7 )
      Move(in := "Datos_maquina".Cinta_en_marcha, out1 => "Mando_driver_cinta")
      Contact( "Q_distancia" )
      R_Coil( "Modo_automatico_DB".Etapa_7 )
      S_Coil( "Modo_automatico_DB".Etapa_8 )
   END_RUNG
   // the same network as SCL:
   IF "Modo_automatico_DB".Etapa_7 THEN "Mando_driver_cinta" := "Datos_maquina".Cinta_en_marcha; END_IF;
   #_w1 := "Modo_automatico_DB".Etapa_7 AND "Q_distancia";
   IF #_w1 THEN
       "Modo_automatico_DB".Etapa_7 := FALSE;
       "Modo_automatico_DB".Etapa_8 := TRUE;
   END_IF;
END_REGION

REGION Network 12: Etapa 8
   // Detener la cinta, cargar tapa
   IF "Modo_automatico_DB".Etapa_8 THEN "Mando_driver_cinta" := "Datos_maquina".Cinta_en_espera; END_IF;
   "IEC_Timer_0_DB_2".TON(IN := "Modo_automatico_DB".Etapa_8, PT := T#2s);
   IF "IEC_Timer_0_DB_2".Q THEN
       "Cargar_tapa_retroceder" := FALSE;
       "Cargar_tapa_avanzar" := TRUE;
   END_IF;
   IF "IEC_Timer_0_DB_2".Q AND "Cargar_tapa_adelante" THEN
       "Modo_automatico_DB".Etapa_8 := FALSE;
       "Modo_automatico_DB".Etapa_9 := TRUE;
   END_IF;
END_REGION

REGION Network 13: Etapa 9
   // Taponar envase
   RUNG wire#powerrail
      Contact( "Modo_automatico_DB".Etapa_9 )
      R_Coil( "Taponador_retroceder" )
      S_Coil( "Taponador_avanzar" )
      Contact( "Taponador_adelante" )
      R_Coil( "Modo_automatico_DB".Etapa_9 )
      S_Coil( "Modo_automatico_DB".Etapa_10 )
   END_RUNG
   // the same network as SCL:
   IF "Modo_automatico_DB".Etapa_9 THEN
       "Taponador_retroceder" := FALSE;
       "Taponador_avanzar" := TRUE;
   END_IF;
   #_w1 := "Modo_automatico_DB".Etapa_9 AND "Taponador_adelante";
   IF #_w1 THEN
       "Modo_automatico_DB".Etapa_9 := FALSE;
       "Modo_automatico_DB".Etapa_10 := TRUE;
   END_IF;
END_REGION

REGION Network 14: Etapa 10
   // Taponadora a posición de reposo 
   // Programar distancia de la cinta hasta la salida